(* Logix 5000 project; controller MV vendor 1 type 14 code 217 rev 31.11; software revision 31.00; part 18 of 53 *)
(* tags used below, declared in another part *)
   CheckTimeMask : INT;
   CWD : CHECKWORD_FLAGS;
   Delphi_Does_Eng_Func : BOOL;
   MC_CH1_R1 : PlantItem;   // CH1_R1
   MC_CH1_R2 : PlantItem;   // CH1_R2
   MC_CH1_R3 : PlantItem;   // CH1_R3
   MC_CH1_R4 : PlantItem;   // CH1_R4
   MC_N255 : INT[255];   // CHECKWORDS Plant item checkword s
   MC_SP_R2_2 : PlantItem;   // SP_R2_2
   MC_SP_R3_1 : PlantItem;   // SP_R3_1
   MC_SP_R5_1 : PlantItem;   // SP_R5_1
   MC_SP_R5_2 : PlantItem;   // SP_R5_2
   MC_SP_R6_1 : PlantItem;   // SP_R6_1
   MC_SP_R6_2 : PlantItem;   // SP_R6_2
   MC_SP_R6_3 : PlantItem;   // SP_R6_3
   MC_SP_R6_4 : PlantItem;   // SP_R6_4
   MC_SP_R6_5 : PlantItem;   // SP_R6_5
   TempChecktime : DINT;
(* MC_Common, continued *)

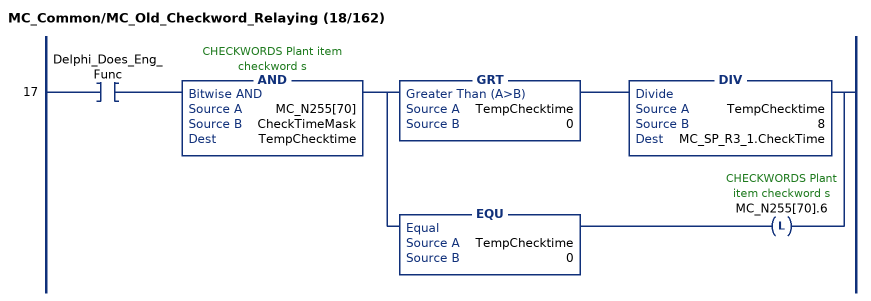
   [picture p288: MC_Common/MC_Old_Checkword_Relaying rungs 17-17]
   17: XIC(Delphi_Does_Eng_Func)AND(MC_N255[70],CheckTimeMask,TempChecktime)[GRT(TempChecktime,0) DIV(TempChecktime,8,MC_SP_R3_1.CheckTime) ,EQU(TempChecktime,0) OTL(MC_N255[70].6) ];
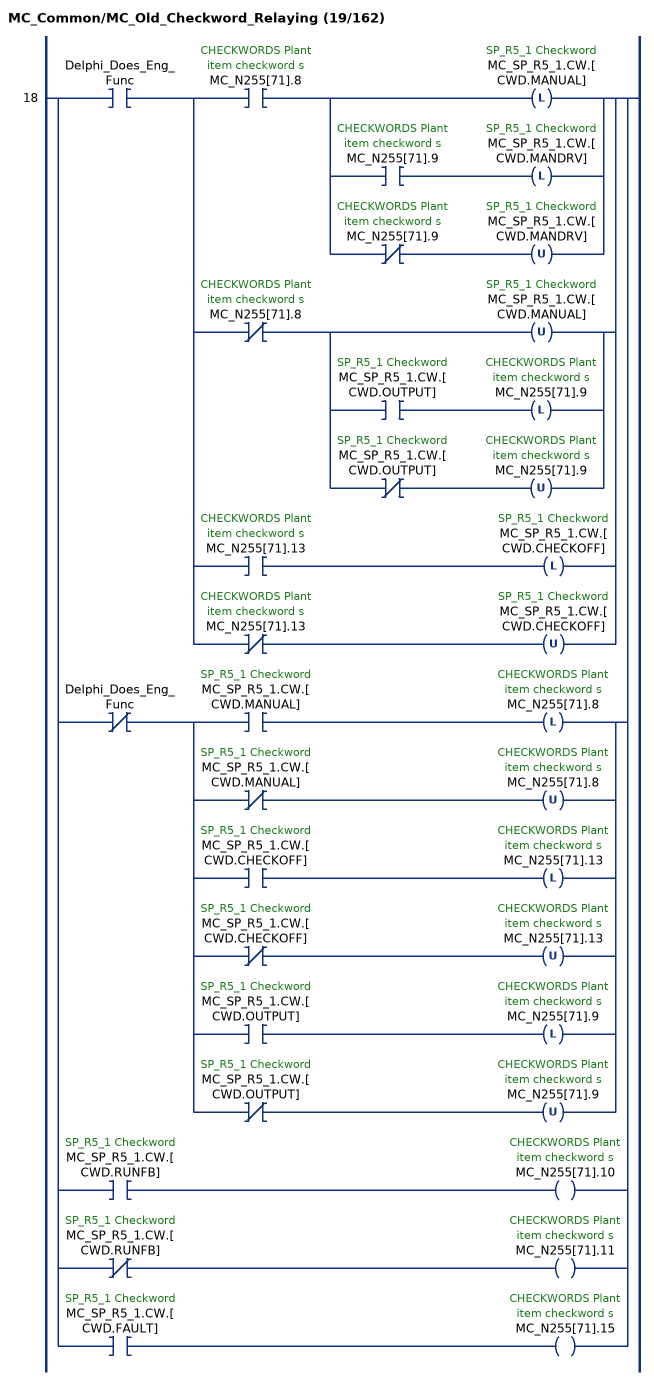
   18: [XIC(Delphi_Does_Eng_Func) [[XIC(MC_N255[71].8) [OTL(MC_SP_R5_1.CW.[CWD.MANUAL]) ,XIC(MC_N255[71].9) OTL(MC_SP_R5_1.CW.[CWD.MANDRV]) ,XIO(MC_N255[71].9) OTU(MC_SP_R5_1.CW.[CWD.MANDRV]) ] ,XIO(MC_N255[71].8) [OTU(MC_SP_R5_1.CW.[CWD.MANUAL]) ,[XIC(MC_SP_R5_1.CW.[CWD.OUTPUT]) OTL(MC_N255[71].9) ,XIO(MC_SP_R5_1.CW.[CWD.OUTPUT]) OTU(MC_N255[71].9) ] ] ] ,[XIC(MC_N255[71].13) OTL(MC_SP_R5_1.CW.[CWD.CHECKOFF]) ,XIO(MC_N255[71].13) OTU(MC_SP_R5_1.CW.[CWD.CHECKOFF]) ] ] ,XIO(Delphi_Does_Eng_Func) [[XIC(MC_SP_R5_1.CW.[CWD.MANUAL]) OTL(MC_N255[71].8) ,XIO(MC_SP_R5_1.CW.[CWD.MANUAL]) OTU(MC_N255[71].8) ] ,[XIC(MC_SP_R5_1.CW.[CWD.CHECKOFF]) OTL(MC_N255[71].13) ,XIO(MC_SP_R5_1.CW.[CWD.CHECKOFF]) OTU(MC_N255[71].13) ] ,[XIC(MC_SP_R5_1.CW.[CWD.OUTPUT]) OTL(MC_N255[71].9) ,XIO(MC_SP_R5_1.CW.[CWD.OUTPUT]) OTU(MC_N255[71].9) ] ] ,XIC(MC_SP_R5_1.CW.[CWD.RUNFB]) OTE(MC_N255[71].10) ,XIO(MC_SP_R5_1.CW.[CWD.RUNFB]) OTE(MC_N255[71].11) ,XIC(MC_SP_R5_1.CW.[CWD.FAULT]) OTE(MC_N255[71].15) ];
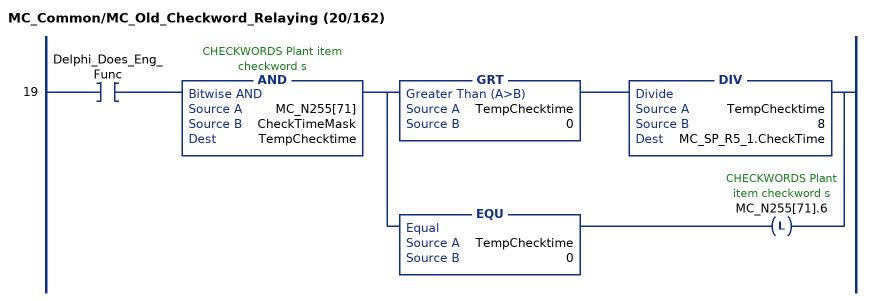
   19: XIC(Delphi_Does_Eng_Func)AND(MC_N255[71],CheckTimeMask,TempChecktime)[GRT(TempChecktime,0) DIV(TempChecktime,8,MC_SP_R5_1.CheckTime) ,EQU(TempChecktime,0) OTL(MC_N255[71].6) ];
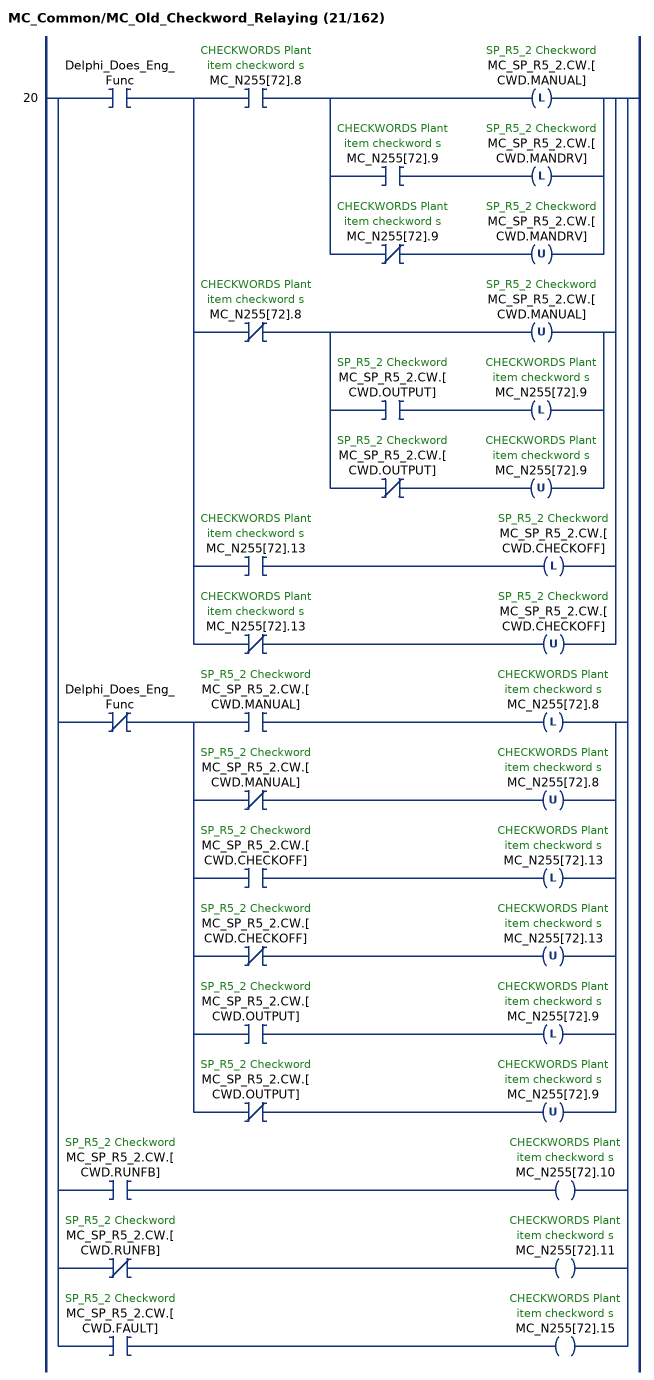
   20: [XIC(Delphi_Does_Eng_Func) [[XIC(MC_N255[72].8) [OTL(MC_SP_R5_2.CW.[CWD.MANUAL]) ,XIC(MC_N255[72].9) OTL(MC_SP_R5_2.CW.[CWD.MANDRV]) ,XIO(MC_N255[72].9) OTU(MC_SP_R5_2.CW.[CWD.MANDRV]) ] ,XIO(MC_N255[72].8) [OTU(MC_SP_R5_2.CW.[CWD.MANUAL]) ,[XIC(MC_SP_R5_2.CW.[CWD.OUTPUT]) OTL(MC_N255[72].9) ,XIO(MC_SP_R5_2.CW.[CWD.OUTPUT]) OTU(MC_N255[72].9) ] ] ] ,[XIC(MC_N255[72].13) OTL(MC_SP_R5_2.CW.[CWD.CHECKOFF]) ,XIO(MC_N255[72].13) OTU(MC_SP_R5_2.CW.[CWD.CHECKOFF]) ] ] ,XIO(Delphi_Does_Eng_Func) [[XIC(MC_SP_R5_2.CW.[CWD.MANUAL]) OTL(MC_N255[72].8) ,XIO(MC_SP_R5_2.CW.[CWD.MANUAL]) OTU(MC_N255[72].8) ] ,[XIC(MC_SP_R5_2.CW.[CWD.CHECKOFF]) OTL(MC_N255[72].13) ,XIO(MC_SP_R5_2.CW.[CWD.CHECKOFF]) OTU(MC_N255[72].13) ] ,[XIC(MC_SP_R5_2.CW.[CWD.OUTPUT]) OTL(MC_N255[72].9) ,XIO(MC_SP_R5_2.CW.[CWD.OUTPUT]) OTU(MC_N255[72].9) ] ] ,XIC(MC_SP_R5_2.CW.[CWD.RUNFB]) OTE(MC_N255[72].10) ,XIO(MC_SP_R5_2.CW.[CWD.RUNFB]) OTE(MC_N255[72].11) ,XIC(MC_SP_R5_2.CW.[CWD.FAULT]) OTE(MC_N255[72].15) ];
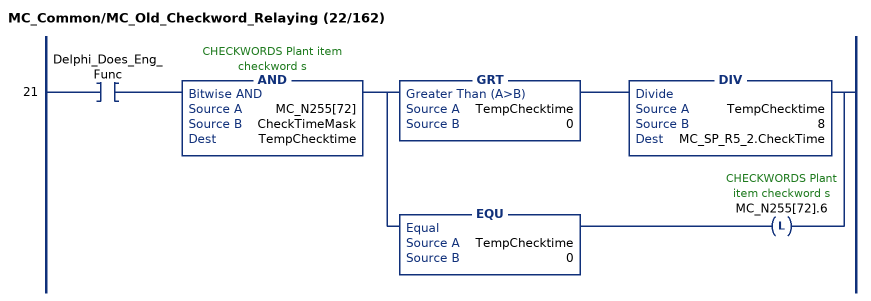
   21: XIC(Delphi_Does_Eng_Func)AND(MC_N255[72],CheckTimeMask,TempChecktime)[GRT(TempChecktime,0) DIV(TempChecktime,8,MC_SP_R5_2.CheckTime) ,EQU(TempChecktime,0) OTL(MC_N255[72].6) ];
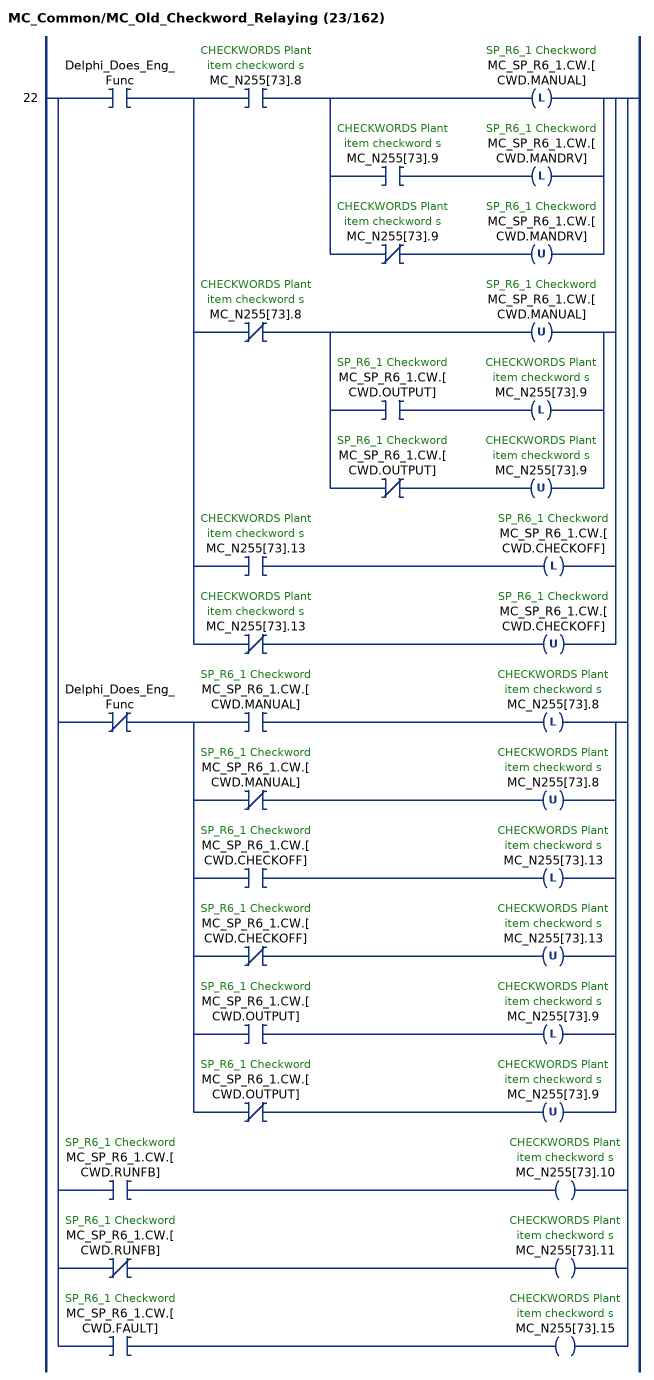
   22: [XIC(Delphi_Does_Eng_Func) [[XIC(MC_N255[73].8) [OTL(MC_SP_R6_1.CW.[CWD.MANUAL]) ,XIC(MC_N255[73].9) OTL(MC_SP_R6_1.CW.[CWD.MANDRV]) ,XIO(MC_N255[73].9) OTU(MC_SP_R6_1.CW.[CWD.MANDRV]) ] ,XIO(MC_N255[73].8) [OTU(MC_SP_R6_1.CW.[CWD.MANUAL]) ,[XIC(MC_SP_R6_1.CW.[CWD.OUTPUT]) OTL(MC_N255[73].9) ,XIO(MC_SP_R6_1.CW.[CWD.OUTPUT]) OTU(MC_N255[73].9) ] ] ] ,[XIC(MC_N255[73].13) OTL(MC_SP_R6_1.CW.[CWD.CHECKOFF]) ,XIO(MC_N255[73].13) OTU(MC_SP_R6_1.CW.[CWD.CHECKOFF]) ] ] ,XIO(Delphi_Does_Eng_Func) [[XIC(MC_SP_R6_1.CW.[CWD.MANUAL]) OTL(MC_N255[73].8) ,XIO(MC_SP_R6_1.CW.[CWD.MANUAL]) OTU(MC_N255[73].8) ] ,[XIC(MC_SP_R6_1.CW.[CWD.CHECKOFF]) OTL(MC_N255[73].13) ,XIO(MC_SP_R6_1.CW.[CWD.CHECKOFF]) OTU(MC_N255[73].13) ] ,[XIC(MC_SP_R6_1.CW.[CWD.OUTPUT]) OTL(MC_N255[73].9) ,XIO(MC_SP_R6_1.CW.[CWD.OUTPUT]) OTU(MC_N255[73].9) ] ] ,XIC(MC_SP_R6_1.CW.[CWD.RUNFB]) OTE(MC_N255[73].10) ,XIO(MC_SP_R6_1.CW.[CWD.RUNFB]) OTE(MC_N255[73].11) ,XIC(MC_SP_R6_1.CW.[CWD.FAULT]) OTE(MC_N255[73].15) ];
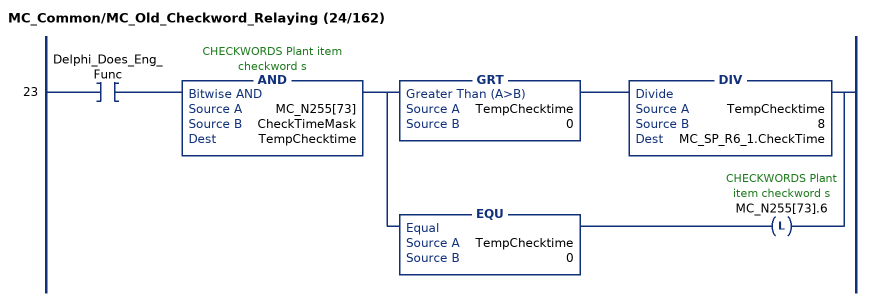
   23: XIC(Delphi_Does_Eng_Func)AND(MC_N255[73],CheckTimeMask,TempChecktime)[GRT(TempChecktime,0) DIV(TempChecktime,8,MC_SP_R6_1.CheckTime) ,EQU(TempChecktime,0) OTL(MC_N255[73].6) ];
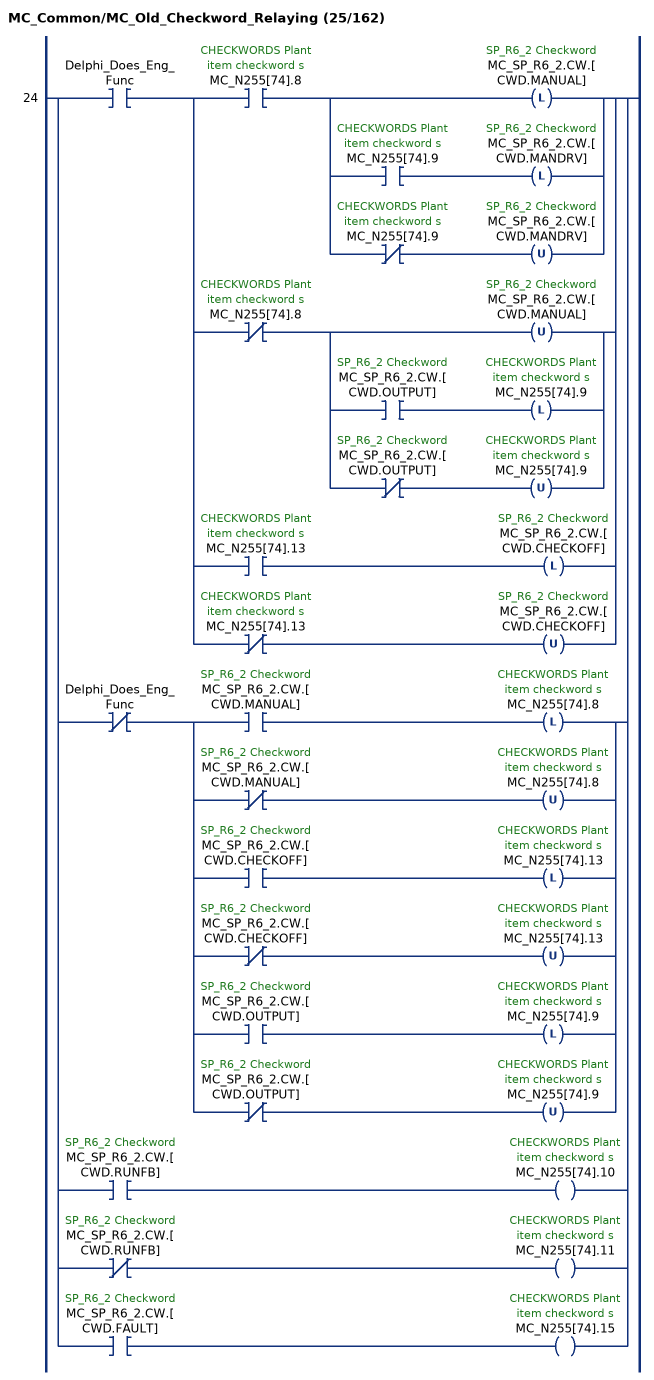
   24: [XIC(Delphi_Does_Eng_Func) [[XIC(MC_N255[74].8) [OTL(MC_SP_R6_2.CW.[CWD.MANUAL]) ,XIC(MC_N255[74].9) OTL(MC_SP_R6_2.CW.[CWD.MANDRV]) ,XIO(MC_N255[74].9) OTU(MC_SP_R6_2.CW.[CWD.MANDRV]) ] ,XIO(MC_N255[74].8) [OTU(MC_SP_R6_2.CW.[CWD.MANUAL]) ,[XIC(MC_SP_R6_2.CW.[CWD.OUTPUT]) OTL(MC_N255[74].9) ,XIO(MC_SP_R6_2.CW.[CWD.OUTPUT]) OTU(MC_N255[74].9) ] ] ] ,[XIC(MC_N255[74].13) OTL(MC_SP_R6_2.CW.[CWD.CHECKOFF]) ,XIO(MC_N255[74].13) OTU(MC_SP_R6_2.CW.[CWD.CHECKOFF]) ] ] ,XIO(Delphi_Does_Eng_Func) [[XIC(MC_SP_R6_2.CW.[CWD.MANUAL]) OTL(MC_N255[74].8) ,XIO(MC_SP_R6_2.CW.[CWD.MANUAL]) OTU(MC_N255[74].8) ] ,[XIC(MC_SP_R6_2.CW.[CWD.CHECKOFF]) OTL(MC_N255[74].13) ,XIO(MC_SP_R6_2.CW.[CWD.CHECKOFF]) OTU(MC_N255[74].13) ] ,[XIC(MC_SP_R6_2.CW.[CWD.OUTPUT]) OTL(MC_N255[74].9) ,XIO(MC_SP_R6_2.CW.[CWD.OUTPUT]) OTU(MC_N255[74].9) ] ] ,XIC(MC_SP_R6_2.CW.[CWD.RUNFB]) OTE(MC_N255[74].10) ,XIO(MC_SP_R6_2.CW.[CWD.RUNFB]) OTE(MC_N255[74].11) ,XIC(MC_SP_R6_2.CW.[CWD.FAULT]) OTE(MC_N255[74].15) ];
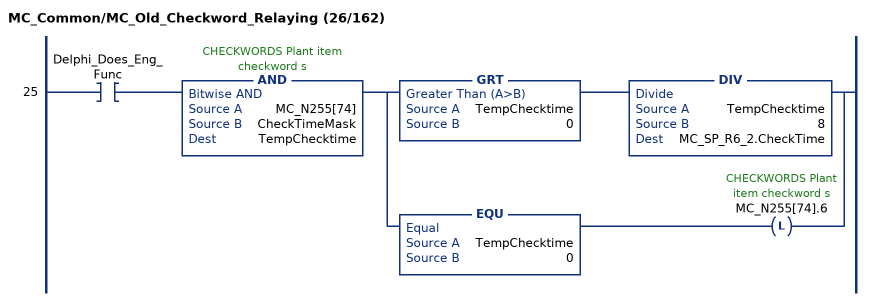
   25: XIC(Delphi_Does_Eng_Func)AND(MC_N255[74],CheckTimeMask,TempChecktime)[GRT(TempChecktime,0) DIV(TempChecktime,8,MC_SP_R6_2.CheckTime) ,EQU(TempChecktime,0) OTL(MC_N255[74].6) ];
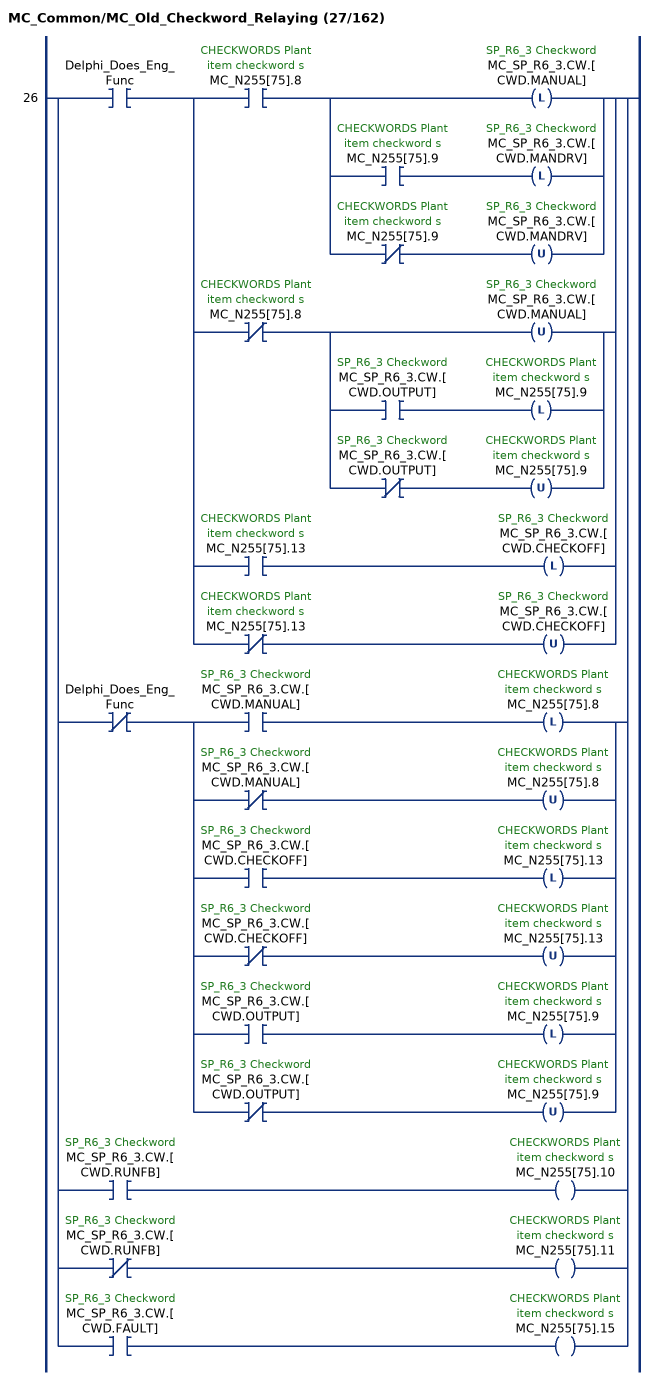
   26: [XIC(Delphi_Does_Eng_Func) [[XIC(MC_N255[75].8) [OTL(MC_SP_R6_3.CW.[CWD.MANUAL]) ,XIC(MC_N255[75].9) OTL(MC_SP_R6_3.CW.[CWD.MANDRV]) ,XIO(MC_N255[75].9) OTU(MC_SP_R6_3.CW.[CWD.MANDRV]) ] ,XIO(MC_N255[75].8) [OTU(MC_SP_R6_3.CW.[CWD.MANUAL]) ,[XIC(MC_SP_R6_3.CW.[CWD.OUTPUT]) OTL(MC_N255[75].9) ,XIO(MC_SP_R6_3.CW.[CWD.OUTPUT]) OTU(MC_N255[75].9) ] ] ] ,[XIC(MC_N255[75].13) OTL(MC_SP_R6_3.CW.[CWD.CHECKOFF]) ,XIO(MC_N255[75].13) OTU(MC_SP_R6_3.CW.[CWD.CHECKOFF]) ] ] ,XIO(Delphi_Does_Eng_Func) [[XIC(MC_SP_R6_3.CW.[CWD.MANUAL]) OTL(MC_N255[75].8) ,XIO(MC_SP_R6_3.CW.[CWD.MANUAL]) OTU(MC_N255[75].8) ] ,[XIC(MC_SP_R6_3.CW.[CWD.CHECKOFF]) OTL(MC_N255[75].13) ,XIO(MC_SP_R6_3.CW.[CWD.CHECKOFF]) OTU(MC_N255[75].13) ] ,[XIC(MC_SP_R6_3.CW.[CWD.OUTPUT]) OTL(MC_N255[75].9) ,XIO(MC_SP_R6_3.CW.[CWD.OUTPUT]) OTU(MC_N255[75].9) ] ] ,XIC(MC_SP_R6_3.CW.[CWD.RUNFB]) OTE(MC_N255[75].10) ,XIO(MC_SP_R6_3.CW.[CWD.RUNFB]) OTE(MC_N255[75].11) ,XIC(MC_SP_R6_3.CW.[CWD.FAULT]) OTE(MC_N255[75].15) ];
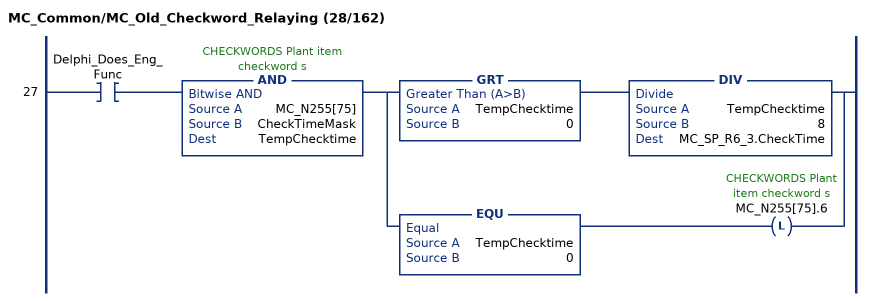
   27: XIC(Delphi_Does_Eng_Func)AND(MC_N255[75],CheckTimeMask,TempChecktime)[GRT(TempChecktime,0) DIV(TempChecktime,8,MC_SP_R6_3.CheckTime) ,EQU(TempChecktime,0) OTL(MC_N255[75].6) ];
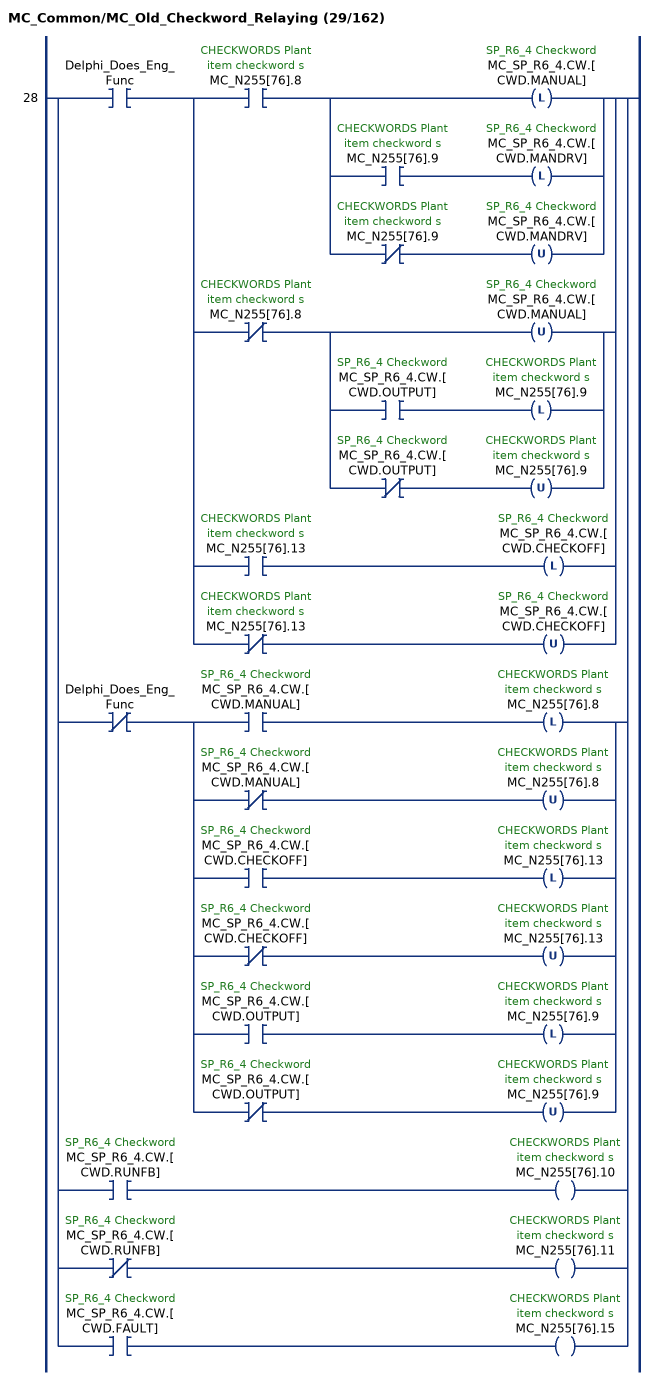
   28: [XIC(Delphi_Does_Eng_Func) [[XIC(MC_N255[76].8) [OTL(MC_SP_R6_4.CW.[CWD.MANUAL]) ,XIC(MC_N255[76].9) OTL(MC_SP_R6_4.CW.[CWD.MANDRV]) ,XIO(MC_N255[76].9) OTU(MC_SP_R6_4.CW.[CWD.MANDRV]) ] ,XIO(MC_N255[76].8) [OTU(MC_SP_R6_4.CW.[CWD.MANUAL]) ,[XIC(MC_SP_R6_4.CW.[CWD.OUTPUT]) OTL(MC_N255[76].9) ,XIO(MC_SP_R6_4.CW.[CWD.OUTPUT]) OTU(MC_N255[76].9) ] ] ] ,[XIC(MC_N255[76].13) OTL(MC_SP_R6_4.CW.[CWD.CHECKOFF]) ,XIO(MC_N255[76].13) OTU(MC_SP_R6_4.CW.[CWD.CHECKOFF]) ] ] ,XIO(Delphi_Does_Eng_Func) [[XIC(MC_SP_R6_4.CW.[CWD.MANUAL]) OTL(MC_N255[76].8) ,XIO(MC_SP_R6_4.CW.[CWD.MANUAL]) OTU(MC_N255[76].8) ] ,[XIC(MC_SP_R6_4.CW.[CWD.CHECKOFF]) OTL(MC_N255[76].13) ,XIO(MC_SP_R6_4.CW.[CWD.CHECKOFF]) OTU(MC_N255[76].13) ] ,[XIC(MC_SP_R6_4.CW.[CWD.OUTPUT]) OTL(MC_N255[76].9) ,XIO(MC_SP_R6_4.CW.[CWD.OUTPUT]) OTU(MC_N255[76].9) ] ] ,XIC(MC_SP_R6_4.CW.[CWD.RUNFB]) OTE(MC_N255[76].10) ,XIO(MC_SP_R6_4.CW.[CWD.RUNFB]) OTE(MC_N255[76].11) ,XIC(MC_SP_R6_4.CW.[CWD.FAULT]) OTE(MC_N255[76].15) ];
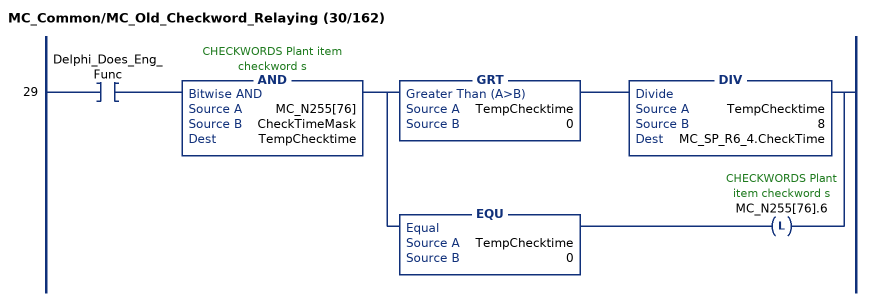
   29: XIC(Delphi_Does_Eng_Func)AND(MC_N255[76],CheckTimeMask,TempChecktime)[GRT(TempChecktime,0) DIV(TempChecktime,8,MC_SP_R6_4.CheckTime) ,EQU(TempChecktime,0) OTL(MC_N255[76].6) ];
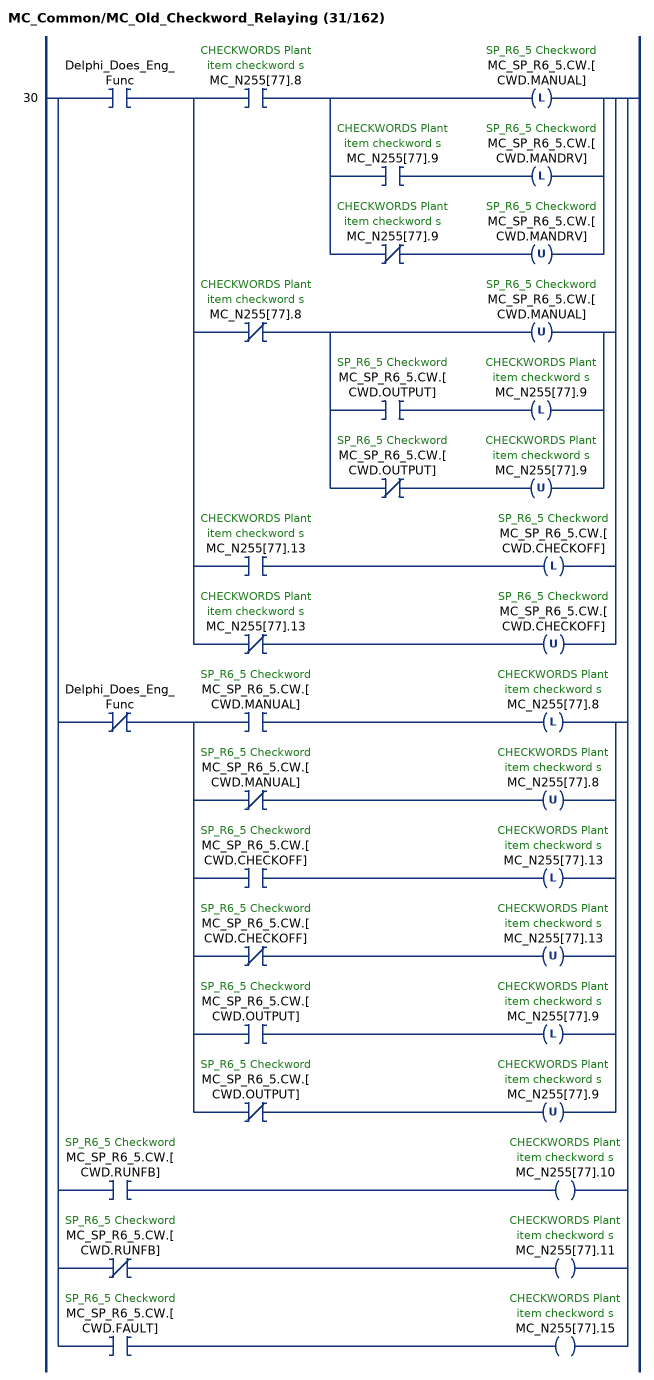
   30: [XIC(Delphi_Does_Eng_Func) [[XIC(MC_N255[77].8) [OTL(MC_SP_R6_5.CW.[CWD.MANUAL]) ,XIC(MC_N255[77].9) OTL(MC_SP_R6_5.CW.[CWD.MANDRV]) ,XIO(MC_N255[77].9) OTU(MC_SP_R6_5.CW.[CWD.MANDRV]) ] ,XIO(MC_N255[77].8) [OTU(MC_SP_R6_5.CW.[CWD.MANUAL]) ,[XIC(MC_SP_R6_5.CW.[CWD.OUTPUT]) OTL(MC_N255[77].9) ,XIO(MC_SP_R6_5.CW.[CWD.OUTPUT]) OTU(MC_N255[77].9) ] ] ] ,[XIC(MC_N255[77].13) OTL(MC_SP_R6_5.CW.[CWD.CHECKOFF]) ,XIO(MC_N255[77].13) OTU(MC_SP_R6_5.CW.[CWD.CHECKOFF]) ] ] ,XIO(Delphi_Does_Eng_Func) [[XIC(MC_SP_R6_5.CW.[CWD.MANUAL]) OTL(MC_N255[77].8) ,XIO(MC_SP_R6_5.CW.[CWD.MANUAL]) OTU(MC_N255[77].8) ] ,[XIC(MC_SP_R6_5.CW.[CWD.CHECKOFF]) OTL(MC_N255[77].13) ,XIO(MC_SP_R6_5.CW.[CWD.CHECKOFF]) OTU(MC_N255[77].13) ] ,[XIC(MC_SP_R6_5.CW.[CWD.OUTPUT]) OTL(MC_N255[77].9) ,XIO(MC_SP_R6_5.CW.[CWD.OUTPUT]) OTU(MC_N255[77].9) ] ] ,XIC(MC_SP_R6_5.CW.[CWD.RUNFB]) OTE(MC_N255[77].10) ,XIO(MC_SP_R6_5.CW.[CWD.RUNFB]) OTE(MC_N255[77].11) ,XIC(MC_SP_R6_5.CW.[CWD.FAULT]) OTE(MC_N255[77].15) ];
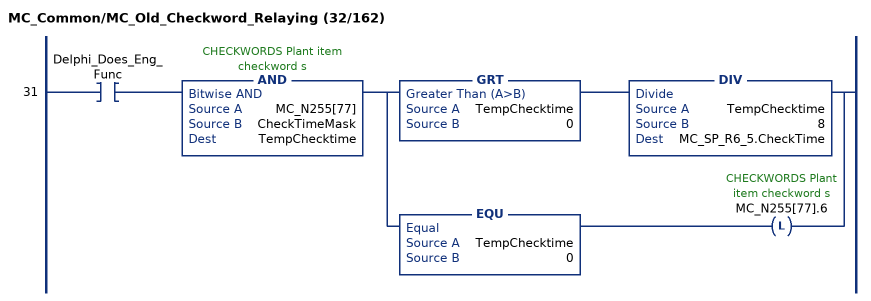
   31: XIC(Delphi_Does_Eng_Func)AND(MC_N255[77],CheckTimeMask,TempChecktime)[GRT(TempChecktime,0) DIV(TempChecktime,8,MC_SP_R6_5.CheckTime) ,EQU(TempChecktime,0) OTL(MC_N255[77].6) ];
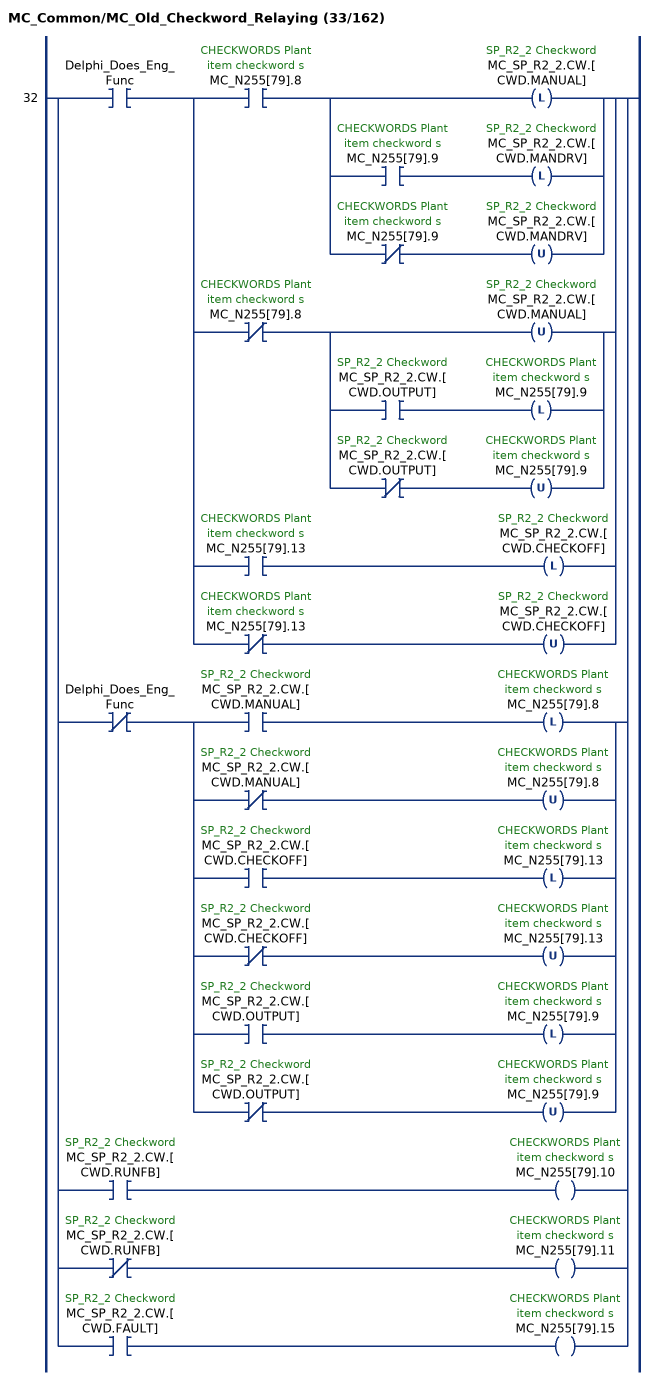
   32: [XIC(Delphi_Does_Eng_Func) [[XIC(MC_N255[79].8) [OTL(MC_SP_R2_2.CW.[CWD.MANUAL]) ,XIC(MC_N255[79].9) OTL(MC_SP_R2_2.CW.[CWD.MANDRV]) ,XIO(MC_N255[79].9) OTU(MC_SP_R2_2.CW.[CWD.MANDRV]) ] ,XIO(MC_N255[79].8) [OTU(MC_SP_R2_2.CW.[CWD.MANUAL]) ,[XIC(MC_SP_R2_2.CW.[CWD.OUTPUT]) OTL(MC_N255[79].9) ,XIO(MC_SP_R2_2.CW.[CWD.OUTPUT]) OTU(MC_N255[79].9) ] ] ] ,[XIC(MC_N255[79].13) OTL(MC_SP_R2_2.CW.[CWD.CHECKOFF]) ,XIO(MC_N255[79].13) OTU(MC_SP_R2_2.CW.[CWD.CHECKOFF]) ] ] ,XIO(Delphi_Does_Eng_Func) [[XIC(MC_SP_R2_2.CW.[CWD.MANUAL]) OTL(MC_N255[79].8) ,XIO(MC_SP_R2_2.CW.[CWD.MANUAL]) OTU(MC_N255[79].8) ] ,[XIC(MC_SP_R2_2.CW.[CWD.CHECKOFF]) OTL(MC_N255[79].13) ,XIO(MC_SP_R2_2.CW.[CWD.CHECKOFF]) OTU(MC_N255[79].13) ] ,[XIC(MC_SP_R2_2.CW.[CWD.OUTPUT]) OTL(MC_N255[79].9) ,XIO(MC_SP_R2_2.CW.[CWD.OUTPUT]) OTU(MC_N255[79].9) ] ] ,XIC(MC_SP_R2_2.CW.[CWD.RUNFB]) OTE(MC_N255[79].10) ,XIO(MC_SP_R2_2.CW.[CWD.RUNFB]) OTE(MC_N255[79].11) ,XIC(MC_SP_R2_2.CW.[CWD.FAULT]) OTE(MC_N255[79].15) ];
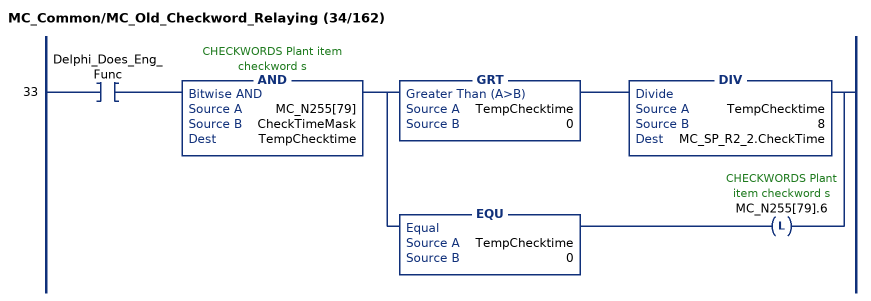
   33: XIC(Delphi_Does_Eng_Func)AND(MC_N255[79],CheckTimeMask,TempChecktime)[GRT(TempChecktime,0) DIV(TempChecktime,8,MC_SP_R2_2.CheckTime) ,EQU(TempChecktime,0) OTL(MC_N255[79].6) ];
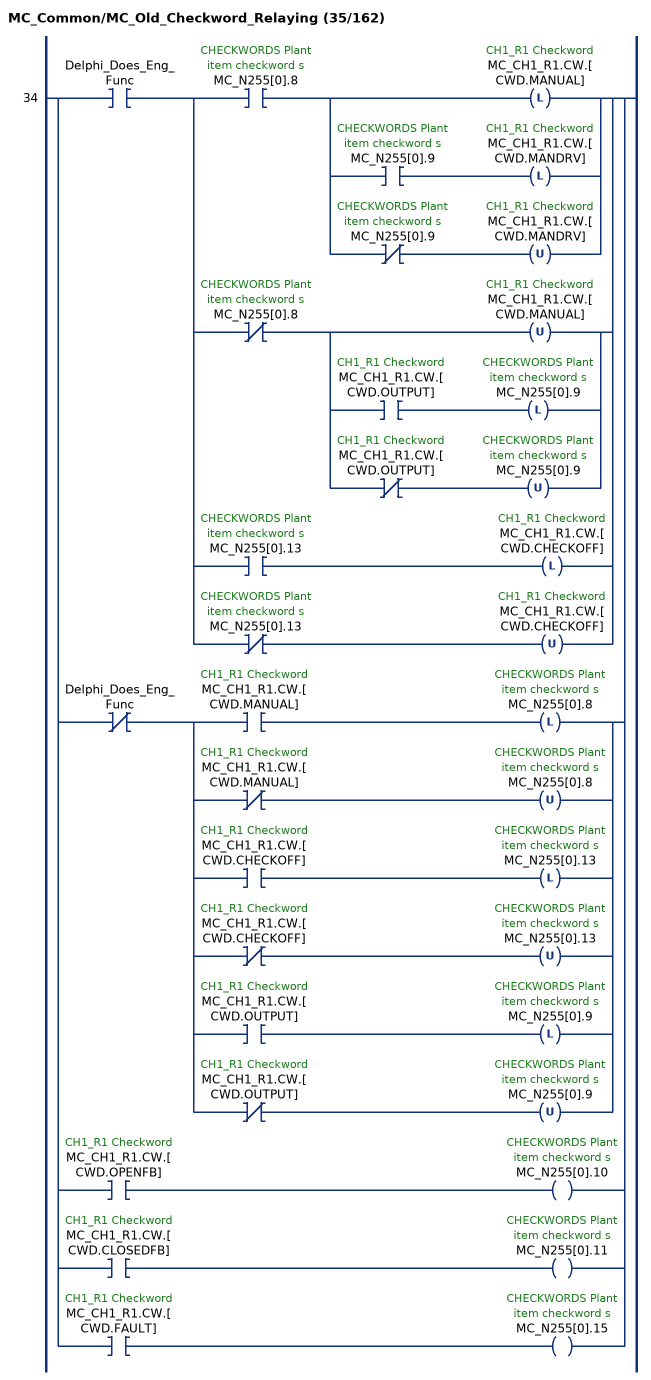
   34: [XIC(Delphi_Does_Eng_Func) [[XIC(MC_N255[0].8) [OTL(MC_CH1_R1.CW.[CWD.MANUAL]) ,XIC(MC_N255[0].9) OTL(MC_CH1_R1.CW.[CWD.MANDRV]) ,XIO(MC_N255[0].9) OTU(MC_CH1_R1.CW.[CWD.MANDRV]) ] ,XIO(MC_N255[0].8) [OTU(MC_CH1_R1.CW.[CWD.MANUAL]) ,[XIC(MC_CH1_R1.CW.[CWD.OUTPUT]) OTL(MC_N255[0].9) ,XIO(MC_CH1_R1.CW.[CWD.OUTPUT]) OTU(MC_N255[0].9) ] ] ] ,[XIC(MC_N255[0].13) OTL(MC_CH1_R1.CW.[CWD.CHECKOFF]) ,XIO(MC_N255[0].13) OTU(MC_CH1_R1.CW.[CWD.CHECKOFF]) ] ] ,XIO(Delphi_Does_Eng_Func) [[XIC(MC_CH1_R1.CW.[CWD.MANUAL]) OTL(MC_N255[0].8) ,XIO(MC_CH1_R1.CW.[CWD.MANUAL]) OTU(MC_N255[0].8) ] ,[XIC(MC_CH1_R1.CW.[CWD.CHECKOFF]) OTL(MC_N255[0].13) ,XIO(MC_CH1_R1.CW.[CWD.CHECKOFF]) OTU(MC_N255[0].13) ] ,[XIC(MC_CH1_R1.CW.[CWD.OUTPUT]) OTL(MC_N255[0].9) ,XIO(MC_CH1_R1.CW.[CWD.OUTPUT]) OTU(MC_N255[0].9) ] ] ,XIC(MC_CH1_R1.CW.[CWD.OPENFB]) OTE(MC_N255[0].10) ,XIC(MC_CH1_R1.CW.[CWD.CLOSEDFB]) OTE(MC_N255[0].11) ,XIC(MC_CH1_R1.CW.[CWD.FAULT]) OTE(MC_N255[0].15) ];
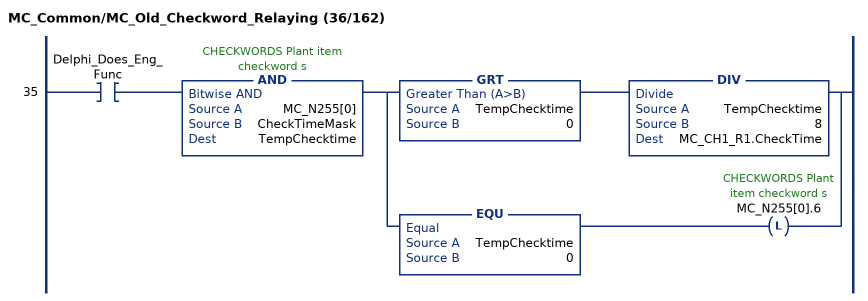
   35: XIC(Delphi_Does_Eng_Func)AND(MC_N255[0],CheckTimeMask,TempChecktime)[GRT(TempChecktime,0) DIV(TempChecktime,8,MC_CH1_R1.CheckTime) ,EQU(TempChecktime,0) OTL(MC_N255[0].6) ];
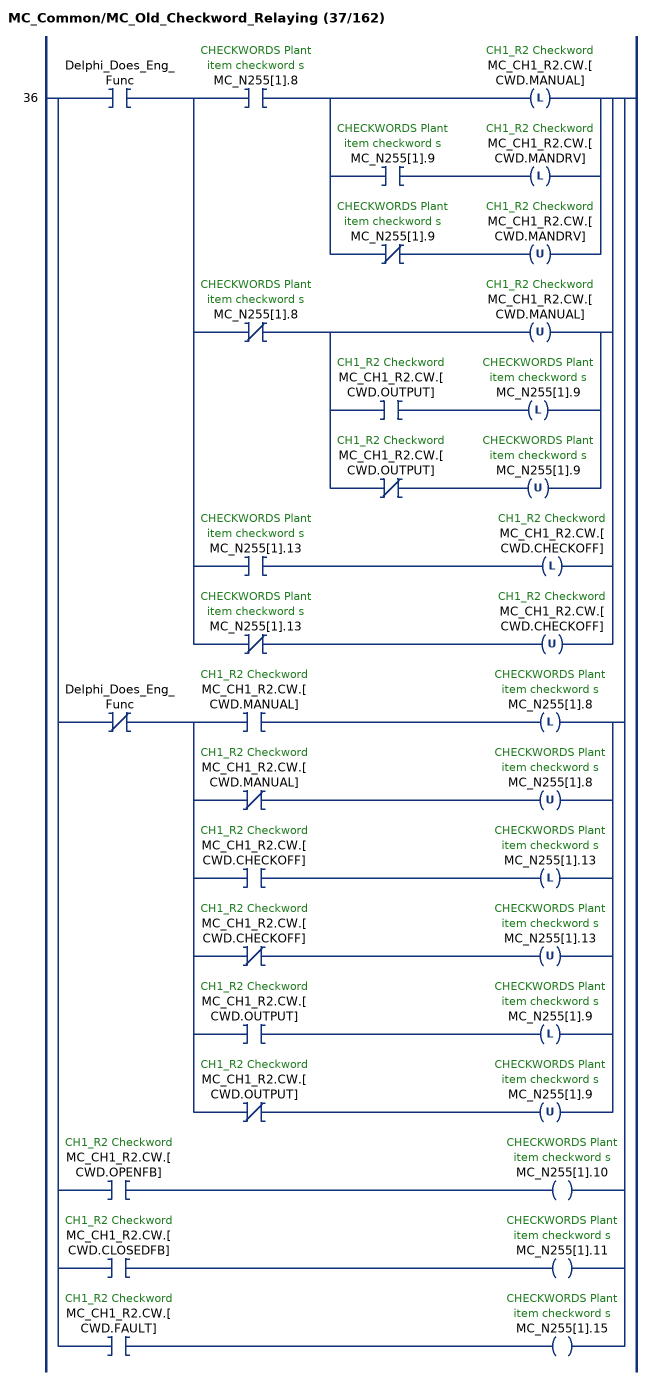
   36: [XIC(Delphi_Does_Eng_Func) [[XIC(MC_N255[1].8) [OTL(MC_CH1_R2.CW.[CWD.MANUAL]) ,XIC(MC_N255[1].9) OTL(MC_CH1_R2.CW.[CWD.MANDRV]) ,XIO(MC_N255[1].9) OTU(MC_CH1_R2.CW.[CWD.MANDRV]) ] ,XIO(MC_N255[1].8) [OTU(MC_CH1_R2.CW.[CWD.MANUAL]) ,[XIC(MC_CH1_R2.CW.[CWD.OUTPUT]) OTL(MC_N255[1].9) ,XIO(MC_CH1_R2.CW.[CWD.OUTPUT]) OTU(MC_N255[1].9) ] ] ] ,[XIC(MC_N255[1].13) OTL(MC_CH1_R2.CW.[CWD.CHECKOFF]) ,XIO(MC_N255[1].13) OTU(MC_CH1_R2.CW.[CWD.CHECKOFF]) ] ] ,XIO(Delphi_Does_Eng_Func) [[XIC(MC_CH1_R2.CW.[CWD.MANUAL]) OTL(MC_N255[1].8) ,XIO(MC_CH1_R2.CW.[CWD.MANUAL]) OTU(MC_N255[1].8) ] ,[XIC(MC_CH1_R2.CW.[CWD.CHECKOFF]) OTL(MC_N255[1].13) ,XIO(MC_CH1_R2.CW.[CWD.CHECKOFF]) OTU(MC_N255[1].13) ] ,[XIC(MC_CH1_R2.CW.[CWD.OUTPUT]) OTL(MC_N255[1].9) ,XIO(MC_CH1_R2.CW.[CWD.OUTPUT]) OTU(MC_N255[1].9) ] ] ,XIC(MC_CH1_R2.CW.[CWD.OPENFB]) OTE(MC_N255[1].10) ,XIC(MC_CH1_R2.CW.[CWD.CLOSEDFB]) OTE(MC_N255[1].11) ,XIC(MC_CH1_R2.CW.[CWD.FAULT]) OTE(MC_N255[1].15) ];
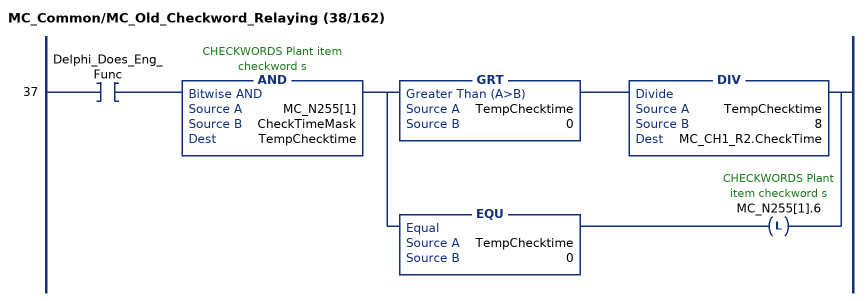
   37: XIC(Delphi_Does_Eng_Func)AND(MC_N255[1],CheckTimeMask,TempChecktime)[GRT(TempChecktime,0) DIV(TempChecktime,8,MC_CH1_R2.CheckTime) ,EQU(TempChecktime,0) OTL(MC_N255[1].6) ];
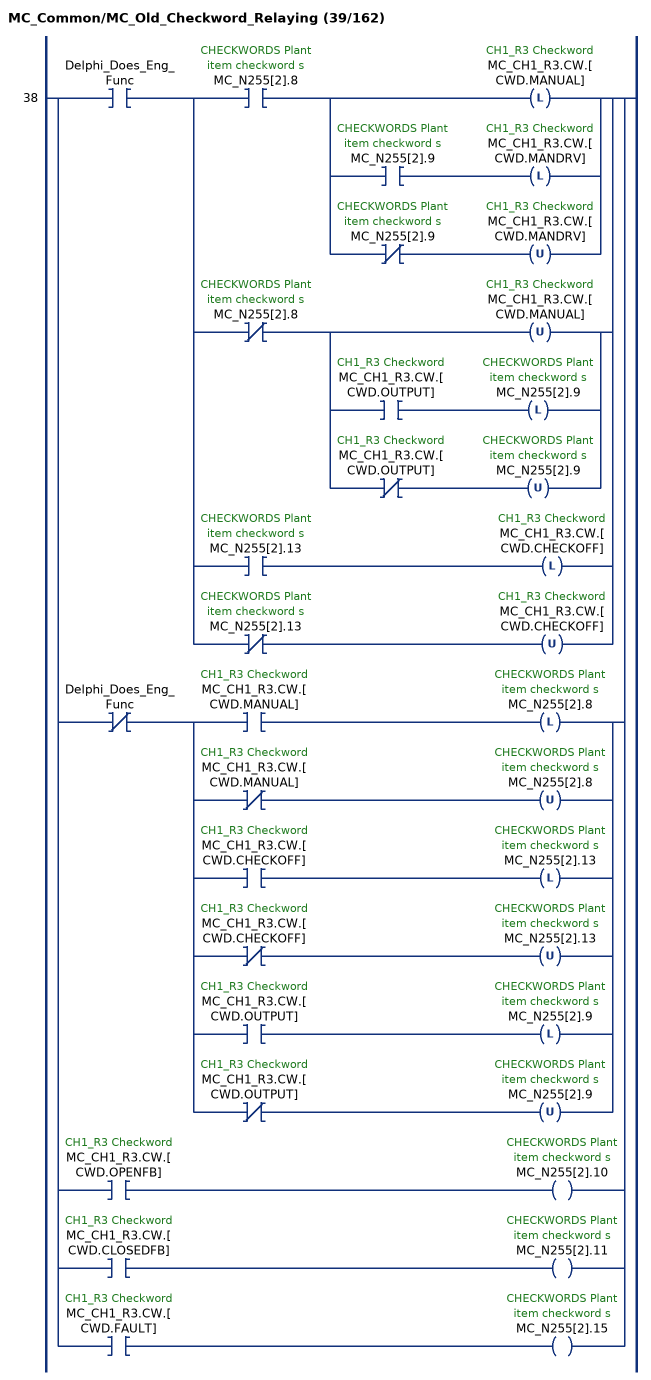
   38: [XIC(Delphi_Does_Eng_Func) [[XIC(MC_N255[2].8) [OTL(MC_CH1_R3.CW.[CWD.MANUAL]) ,XIC(MC_N255[2].9) OTL(MC_CH1_R3.CW.[CWD.MANDRV]) ,XIO(MC_N255[2].9) OTU(MC_CH1_R3.CW.[CWD.MANDRV]) ] ,XIO(MC_N255[2].8) [OTU(MC_CH1_R3.CW.[CWD.MANUAL]) ,[XIC(MC_CH1_R3.CW.[CWD.OUTPUT]) OTL(MC_N255[2].9) ,XIO(MC_CH1_R3.CW.[CWD.OUTPUT]) OTU(MC_N255[2].9) ] ] ] ,[XIC(MC_N255[2].13) OTL(MC_CH1_R3.CW.[CWD.CHECKOFF]) ,XIO(MC_N255[2].13) OTU(MC_CH1_R3.CW.[CWD.CHECKOFF]) ] ] ,XIO(Delphi_Does_Eng_Func) [[XIC(MC_CH1_R3.CW.[CWD.MANUAL]) OTL(MC_N255[2].8) ,XIO(MC_CH1_R3.CW.[CWD.MANUAL]) OTU(MC_N255[2].8) ] ,[XIC(MC_CH1_R3.CW.[CWD.CHECKOFF]) OTL(MC_N255[2].13) ,XIO(MC_CH1_R3.CW.[CWD.CHECKOFF]) OTU(MC_N255[2].13) ] ,[XIC(MC_CH1_R3.CW.[CWD.OUTPUT]) OTL(MC_N255[2].9) ,XIO(MC_CH1_R3.CW.[CWD.OUTPUT]) OTU(MC_N255[2].9) ] ] ,XIC(MC_CH1_R3.CW.[CWD.OPENFB]) OTE(MC_N255[2].10) ,XIC(MC_CH1_R3.CW.[CWD.CLOSEDFB]) OTE(MC_N255[2].11) ,XIC(MC_CH1_R3.CW.[CWD.FAULT]) OTE(MC_N255[2].15) ];
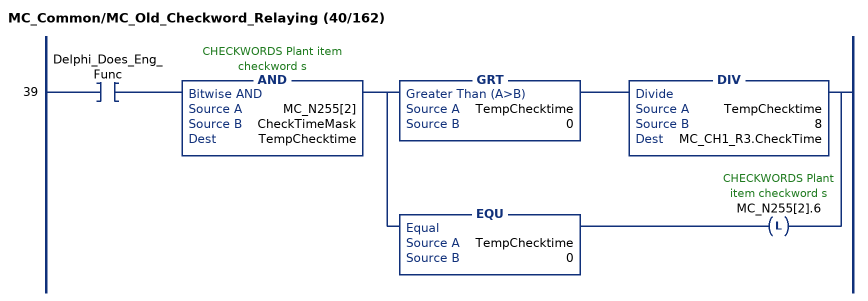
   39: XIC(Delphi_Does_Eng_Func)AND(MC_N255[2],CheckTimeMask,TempChecktime)[GRT(TempChecktime,0) DIV(TempChecktime,8,MC_CH1_R3.CheckTime) ,EQU(TempChecktime,0) OTL(MC_N255[2].6) ];
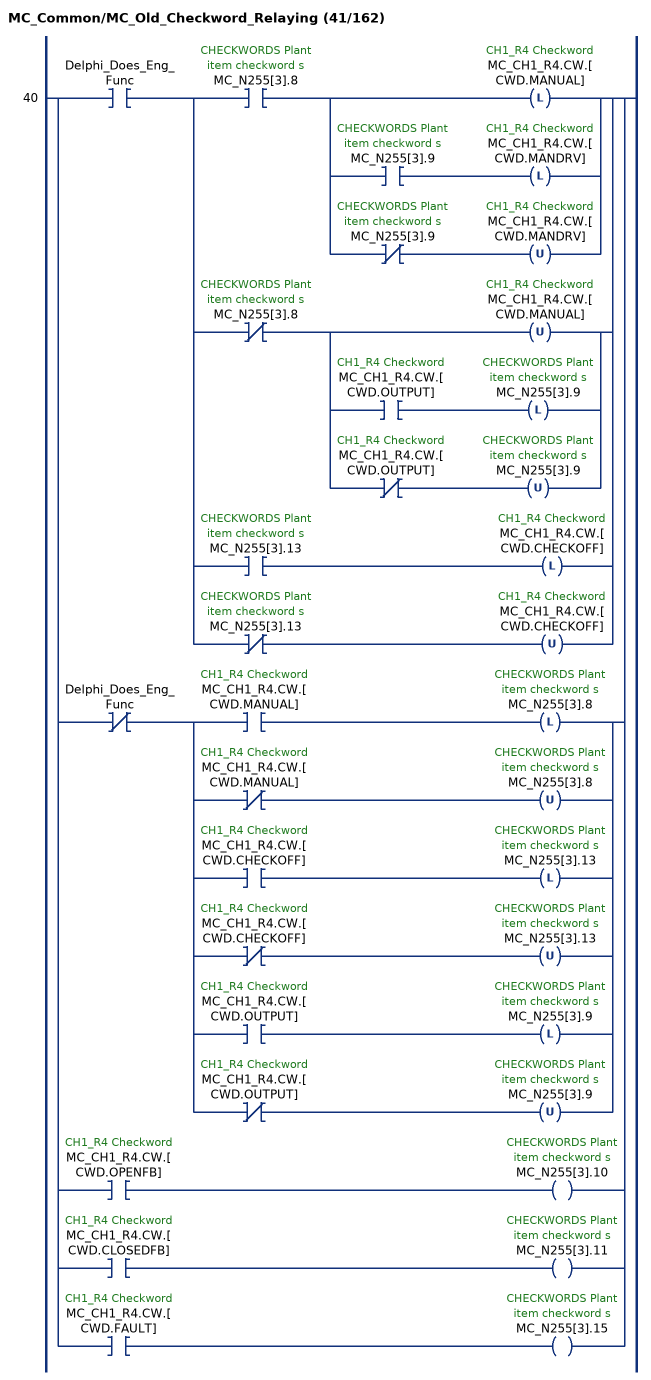
   40: [XIC(Delphi_Does_Eng_Func) [[XIC(MC_N255[3].8) [OTL(MC_CH1_R4.CW.[CWD.MANUAL]) ,XIC(MC_N255[3].9) OTL(MC_CH1_R4.CW.[CWD.MANDRV]) ,XIO(MC_N255[3].9) OTU(MC_CH1_R4.CW.[CWD.MANDRV]) ] ,XIO(MC_N255[3].8) [OTU(MC_CH1_R4.CW.[CWD.MANUAL]) ,[XIC(MC_CH1_R4.CW.[CWD.OUTPUT]) OTL(MC_N255[3].9) ,XIO(MC_CH1_R4.CW.[CWD.OUTPUT]) OTU(MC_N255[3].9) ] ] ] ,[XIC(MC_N255[3].13) OTL(MC_CH1_R4.CW.[CWD.CHECKOFF]) ,XIO(MC_N255[3].13) OTU(MC_CH1_R4.CW.[CWD.CHECKOFF]) ] ] ,XIO(Delphi_Does_Eng_Func) [[XIC(MC_CH1_R4.CW.[CWD.MANUAL]) OTL(MC_N255[3].8) ,XIO(MC_CH1_R4.CW.[CWD.MANUAL]) OTU(MC_N255[3].8) ] ,[XIC(MC_CH1_R4.CW.[CWD.CHECKOFF]) OTL(MC_N255[3].13) ,XIO(MC_CH1_R4.CW.[CWD.CHECKOFF]) OTU(MC_N255[3].13) ] ,[XIC(MC_CH1_R4.CW.[CWD.OUTPUT]) OTL(MC_N255[3].9) ,XIO(MC_CH1_R4.CW.[CWD.OUTPUT]) OTU(MC_N255[3].9) ] ] ,XIC(MC_CH1_R4.CW.[CWD.OPENFB]) OTE(MC_N255[3].10) ,XIC(MC_CH1_R4.CW.[CWD.CLOSEDFB]) OTE(MC_N255[3].11) ,XIC(MC_CH1_R4.CW.[CWD.FAULT]) OTE(MC_N255[3].15) ];
